(* Logix 5000 project; controller PLC_MCC1300_75F1 vendor 1 type 14 code 166 rev 32.11; software revision 32.04; part 10 of 83 *)

        [35]   // PEG SAMPLE Trailedge Positioning Timer Preset [sec x 100]
        [4].7   // Stress Sample one shot for new LE at Conv 6 Resync Zone
        [6].9   // 400 Deck Conveyor 9 Operate at Trim speed
        [20].3   // STRESS SAMPLE Stop Conv 8 for Sample Positioning
        [32]   // PEG SAMPLE Trailedge Stopping Setpoint [inches x 10]
        [7].8   // PEG SAMPLE Lead-Cap Runout In Progress (Stop Conv 9)
        [50]   // PEG SAMPLE Trailedge Stopping Setpoint [inches x 10]
        [11]   // Sample/Peg CAP Length in Inches
        [7].7   // Sample/Peg Stop Conv 9 When next CAP Arrives
        [37]   // PEG SAMPLE TE Stopping Setpoint for Glass <> 60 In [inches x 10]
        [90]   // PEG SAMPLE Trailedge Stopping(2100in/min) Setpoint [inches x 10]
        [10]   // Sample/Peg CAP Length + Trailedge Position in Zones
        [41]   // 400 DECK Decel Distance for Current Trim Speed [in]
        [2]   // 400 DECK CAP Length of Current Cap [64ths]
        [8]   // Sample/Peg Transfer State Machine
        [14]   // PEG SAMPLE Minimum Gap + Cap Value for LCR [inches / 2]
        [42]   // 400 DECK CAP Length Divided by 2 for Current Piece [in]
        [5].8   // 400 Deck
        [20].2   // Conveyor 7 Leadedge Detected
        [7].2   // Queue Conv 4 Leadedge Detected
        [20].1   // Conveyor 6 Trailedge Detected
        [7].1   // Queue Conv 4 Trailedge Detected
        [0]   // 400 Deck State Variable
        [45]   // 400 Deck Host ID
        [5].9   // 400 Deck
        [25]   // Heavy Glass Sample Cap ID
        [31]   // PEG SAMPLE Decel Distance at Current Speed for Positioning Calc. [in x 10]
        [4].0   // 400 Deck One shot!
   N98 : DINT[40] := ([0] := 12767, [1] := -2664, [5] := 241, [6] := 245, [7] := 244, [8] := 243, [9] := 230, [10] := 232, [11] := 237, [12] := 239);
   O : INT[128] := ([5] := 2#0000_1111_1111_1111, [8] := 2#0000_1000_0000_0000, [9] := 2#0010_0000_0000_1000, [17] := 2#0000_0000_0000_1000, [21] := 2#1111_1100_0000_1000, [23] := 2#0000_0000_0000_0011, [27] := 2#0001_0000_0000_0010, [29] := 2#0001_0000_0000_0010, [30] := 2#0010_0100_0011_1111, [31] := 2#0001_0000_0000_0010, [34] := 2#0000_0000_0000_0110, [38] := 2#0000_0000_0110_0011, [41] := 2#0000_0001_0000_0000, [42] := 2#0000_0000_0000_0100, [46] := 2#0000_0000_0000_0100, [50] := 2#0000_0000_0000_0011, [62] := 2#0000_0000_0000_0011, [66] := 2#0000_0000_0000_0100, [70] := 2#0000_0000_0000_0100, [74] := 2#1000_0100_1100_0011, [78] := 2#0000_0000_0000_0010, [80] := 2#0000_0000_0111_1011, [81] := 2#0000_0010_0100_0000, [82] := 2#0000_0000_0100_0011, [83] := 2#0000_0001_0100_0001, [84] := 2#0000_0001_0100_0001, [85] := 2#0001_0001_0100_0010, [86] := 2#0000_0001_0100_0001, [87] := 2#0001_0000_0000_0010, [89] := 2#0001_0000_0000_0010, [91] := 2#0001_0000_0000_0010, [92] := 2#0000_1001_1100_1010, [93] := 2#0011_0000_0000_0010, [95] := 2#0011_0000_0000_0010, [96] := 2#0000_0000_0000_0011, [97] := 2#0011_0000_0000_0010, [99] := 2#0011_0000_0000_0010, [101] := 2#0011_0001_1100_0010, [103] := 2#0011_0000_0000_0010, [105] := 2#0011_0000_0000_0010, [107] := 2#0011_0000_0000_0010, [109] := 2#0011_0000_0000_0010, [111] := 2#0011_0000_0000_0010, [113] := 2#0011_0000_0000_0010, [115] := 2#0011_0000_0000_0010, [117] := 2#0011_0000_0000_0010, [119] := 2#0011_0000_0000_0010, [121] := 2#0000_0000_1000_0100, [123] := 2#0000_1000_0000_0000);
        [113].8   // VMCC M2 Speed zone 11 Accel Rate Select 1 * M2CM11S
        [113].9   // VMCC M2 Speed zone 11 Accel Rate Select 2 * M2CM11S
        [111].9   // VMCC M2 Speed zone 10 Accel Rate Select 2 * M2CM10N
        [113].10   // VMCC M2 Speed zone 11 Decel Rate Select 1 * M2CM11S
        [103].11   // VMCC M2 Speed zone 8 Decel Rate Select 2 * M2CM8N
        [105].10   // VMCC M2 Speed zone 9 Decel Rate Select 1 * M2CM9S
        [105].11   // VMCC M2 Speed zone 9 Decel Rate Select 2 * M2CM9S
        [107].10   // VMCC M2 Speed zone 9 Decel Rate Select 1 * M2CM9N
        [107].11   // VMCC M2 Speed zone 9 Decel Rate Select 2 * M2CM9N
        [101].2   // VMCC M2 Speed zone 8 Jog * M2CM8S
        [117].6   // VMCC M2 Speed zone 12 Local Control Reques * M2CM12S
        [115].10   // VMCC M2 Speed zone 11 Decel Rate Select 1 * M2CM11N
        [119].4   // VMCC M2 Speed zone 12 Direction Select 1 * M2CM12N
        [119].5   // VMCC M2 Speed zone 12 Direction Select 2 * M2CM12N
        [103].2   // VMCC M2 Speed zone 8 Jog * M2CM8N
        [105].2   // VMCC M2 Speed zone 9 Jog * M2CM9S
        [119].9   // VMCC M2 Speed zone 12 Accel Rate Select 2 * M2CM12N
        [121]   // M2 -->> MB Copy mainline crusher status bits from M2 to MB
        [117].8   // VMCC M2 Speed zone 12 Accel Rate Select 1 * M2CM12S
        [123].2   // M2 -->> MB Trim deck Drive system Critical Failure
        [123].5   // M2 -->> MB Mainline Drive system Critical Failure
        [115].8   // VMCC M2 Speed zone 11 Accel Rate Select 1 * M2CM11N
        [101].3   // VMCC M2 Speed zone 8 Clear Fault * M2CM8S
        [107].2   // VMCC M2 Speed zone 9 Jog * M2CM9N
        [123].11   // M2 -->> MB Drive running M2CM01
        [123].3   // M2 -->> MB Trim deck Drive fault
        [25].3   // ROCKWELL CAPPER Disable auto y-cut bar 4
        [27].0   // VMCC M2 Speed zone 1 Stop * M2CM01
        [5].9   // VMCC M2 Speed zone 10 Foward * 2CM10
        [6].0   // VMCC M2 Speed zone 1 Reverse * 2CM01
        [6].1   // VMCC M2 Speed zone 2 Reverse * 2CM02
        [6].2   // VMCC M2 Speed zone 3 Reverse * 2CM03
        [6].3   // VMCC M2 Speed zone 4 Reverse * 2CM04
        [109].2   // VMCC M2 Speed zone 10 Jog * M2CM10S
        [111].2   // VMCC M2 Speed zone 10 Jog * M2CM10N
        [124].0   // M2 -->> MB Leg 4 Is In Sleep Mode
        [103].3   // VMCC M2 Speed zone 8 Clear Fault * M2CM8N
        [6].4   // VMCC M2 Speed zone 5 Reverse * 2CM05
        [124].1   // M2 -->> MB Leg 5 Is In Sleep Mode
        [6].5   // VMCC M2 Speed zone 6 Reverse * 2CM06
        [123].8   // M2 -->> MB SPARE
        [10].10   // VMCC M2 SPARE
        [10].11   // VMCC M2 SPARE
        [123].9   // M2 -->> MB SPARE
        [20].8   // VMCC TD Trim knocker Speed select 2
        [124].4   // M2-->MB VISION SYS Rejected Plate Alarm Horn
        [19].2   // VMCC TD Trim Zone 1 North knocker Adjust motor
        [105].3   // VMCC M2 Speed zone 9 Clear Fault * M2CM9S
        [113].2   // VMCC M2 Speed zone 11 Jog * M2CM11S
        [107].3   // VMCC M2 Speed zone 9 Clear Fault * M2CM9N
        [123].13   // M2 -->> MB Crush-all Selector sw. Status
        [20].9   // VMCC TD Trim deck Speed select 2 North side
        [101].12   // VMCC M2 Speed zone 8 Speed Select 1 * M2CM8S
        [42].5   // RELIANCE CAPPING SYSTEM Tracking window Lamp
        [19].3   // VMCC TD Trim Zone 1 South knocker Adjust motor
        [70].5   // RELIANCE CAPPING SYSTEM Tracking window Lamp
        [115].2   // VMCC M2 Speed zone 11 Jog * M2CM11N
        [19].4   // VMCC TD Trim Zone 2 North knocker Adjust motor
        [19].5   // VMCC TD Trim Zone 2 South knocker Adjust motor
        [27].3   // VMCC M2 Speed zone 1 Clear Fault * M2CM01
        [7].10   // VMCC M2 Speed zone 11 Speed Select 2 * 2CM11
        [22].2   // VMCC TD Trim Zone 1 North trim Adjust motor
        [22].3   // VMCC TD Trim Zone 1 South trim Adjust motor
        [117].9   // VMCC M2 Speed zone 12 Accel Rate Select 2 * M2CM12S
        [74].13   // BENCHBOARD SPARE
        [101].13   // VMCC M2 Speed zone 8 Speed Select 2 * M2CM8S
        [109].10   // VMCC M2 Speed zone 10 Decel Rate Select 1 * M2CM10S
        [109].11   // VMCC M2 Speed zone 10 Decel Rate Select 2 * M2CM10S
        [109].6   // VMCC M2 Speed zone 10 Local Control Reques * M2CM10S
        [109].8   // VMCC M2 Speed zone 10 Accel Rate Select 1 * M2CM10S
        [25].4   // ROCKWELL CAPPER Disable auto y-cut bar 3
        [10].12   // VMCC M2 SPARE
        [10].13   // VMCC M2 SPARE
        [10].14   // VMCC M2 SPARE
        [10].15   // VMCC M2 SPARE
        [19].12   // VMCC TD SPARE
        [19].13   // VMCC TD SPARE
        [19].14   // VMCC TD SPARE
        [19].15   // VMCC TD SPARE
        [101].0   // VMCC M2 Speed zone 8 Stop * M2CM8S
        [19].6   // VMCC TD Trim Zone 3 North knocker Adjust motor
        [125]   // MB -->> M2 Host comp. Reliance Crossbreaks Disable Ycuts
        [119].6   // VMCC M2 Speed zone 12 Local Control Reques * M2CM12N
        [109].0   // VMCC M2 Speed zone 10 Stop * M2CM10S
        [111].0   // VMCC M2 Speed zone 10 Stop * M2CM10N
        [113].0   // VMCC M2 Speed zone 11 Stop * M2CM11S
        [115].0   // VMCC M2 Speed zone 11 Stop * M2CM11N
        [42].2   // PANEL TD-CS2N North Trim knocker #2 Lower
        [46].2   // PANEL TD-CS3N North Trim knocker #3 Lower
        [50].2   // PANEL TD-CS4N North Trim knocker #4 Lower
        [55].2   // PANEL TD-CS5N North Trim knocker #5 Lower
        [62].2   // PANEL TD-CS4S South Trim knocker #4 Lower
        [66].2   // PANEL TD-CS3S South Trim knocker #3 Lower
        [70].2   // PANEL TD-CS2S South Trim knocker #2 Lower
        [7].0   // VMCC M2 Speed zone 1 Speed Select 2 * 2CM01
        [7].1   // VMCC M2 Speed zone 2 Speed Select 2 * 2CM02
        [7].2   // VMCC M2 Speed zone 3 Speed Select 2 * 2CM03
        [7].3   // VMCC M2 Speed zone 4 Speed Select 2 * 2CM04
        [7].4   // VMCC M2 Speed zone 5 Speed Select 2 * 2CM05
        [7].5   // VMCC M2 Speed zone 6 Speed Select 2 * 2CM06
        [7].6   // VMCC M2 Speed zone 7 Speed Select 2 * 2CM07
        [7].7   // VMCC M2 Speed zone 8 Speed Select 2 * 2CM08
        [7].8   // VMCC M2 Speed zone 9 Speed Select 2 * 2CM09
        [85].3   // VMCC M2 Speed zone 4 Clear Fault * M2CM4S
        [87].3   // VMCC M2 Speed zone 4 Clear Fault * M2CM4N
        [22].0   // VMCC TD Krurl drop North trim Adjust motor
        [89].3   // VMCC M2 Speed zone 5 Clear Fault * M2CM5S
        [8].0   // VMCC M2 Speed zone 1 Speed Select 1 * 2CM01
        [8].1   // VMCC M2 Speed zone 2 Speed Select 1 * 2CM02
        [8].2   // VMCC M2 Speed zone 3 Speed Select 1 * 2CM03
        [8].3   // VMCC M2 Speed zone 4 Speed Select 1 * 2CM04
        [8].4   // VMCC M2 Speed zone 5 Speed Select 1 * 2CM05
        [8].5   // VMCC M2 Speed zone 6 Speed Select 1 * 2CM06
        [8].6   // VMCC M2 Speed zone 7 Speed Select 1 * 2CM07
        [8].7   // VMCC M2 Speed zone 8 Speed Select 1 * 2CM08
        [22].1   // VMCC TD Krurl drop South trim Adjust motor
        [25].1   // ROCKWELL CAPPER Disable manual y-cut bar 2
        [8].8   // VMCC M2 Speed zone 9 Speed Select 1 * 2CM09
        [25].5   // ROCKWELL CAPPER Disable auto y-cut bar 2
        [103].0   // VMCC M2 Speed zone 8 Stop * M2CM8N
        [117].0   // VMCC M2 Speed zone 12 Stop * M2CM12S
        [119].0   // VMCC M2 Speed zone 12 Stop * M2CM12N
        [105].0   // VMCC M2 Speed zone 9 Stop * M2CM9S
        [115].11   // VMCC M2 Speed zone 11 Decel Rate Select 2 * M2CM11N
        [91].3   // VMCC M2 Speed zone 5 Clear Fault * M2CM5N
        [117].2   // VMCC M2 Speed zone 12 Jog * M2CM12S
        [119].2   // VMCC M2 Speed zone 12 Jog * M2CM12N
        [123].14   // M2 -->> MB Leg 2 Is In Sleep Mode
        [123].15   // M2 -->> MB Leg 3 Is In Sleep Mode
        [22].4   // VMCC TD Trim Zone 2 North trim Adjust motor
        [20].12   // VMCC TD Trim knocker Speed select 1
        [6].10   // VMCC M2 Speed zone 11 Reverse * 2CM11
        [6].11   // VMCC M2 Speed zone 12 Reverse * 2CM12
        [9].2   // VMCC M2 SPARE
        [123].10   // M2 -->> MB SPARE
        [10].0   // VMCC M2 SPARE
        [22].5   // VMCC TD Trim Zone 2 South trim Adjust motor
        [22].6   // VMCC TD Trim Zone 3 North trim Adjust motor
        [101].14   // VMCC M2 Speed zone 8 Speed Select 3 * M2CM8S
        [103].12   // VMCC M2 Speed zone 8 Speed Select 1 * M2CM8N
        [8].10   // VMCC M2 Speed zone 11 Speed Select 1 * 2CM11
        [19].7   // VMCC TD Trim Zone 3 South knocker Adjust motor
        [8].11   // VMCC M2 Speed zone 12 Speed Select 1 * 2CM12
        [103].13   // VMCC M2 Speed zone 8 Speed Select 2 * M2CM8N
        [19]   // TRIM KNOCKERS Contactors used For drive to Knocker adj Motors
        [119].8   // VMCC M2 Speed zone 12 Accel Rate Select 1 * M2CM12N
        [22].7   // VMCC TD Trim Zone 3 South trim Adjust motor
        [22].8   // VMCC TD Trim Zone 4 North trim Adjust motor
        [103].14   // VMCC M2 Speed zone 8 Speed Select 3 * M2CM8N
        [105].12   // VMCC M2 Speed zone 9 Speed Select 1 * M2CM9S
        [93].3   // VMCC M2 Speed zone 6 Clear Fault * M2CM6S
        [22].9   // VMCC TD Trim Zone 4 South trim Adjust motor
        [27].1   // VMCC M2 Speed zone 1 Forward/start * M2CM01
        [19].8   // VMCC TD Trim Zone 4 North knocker Adjust motor
        [105].13   // VMCC M2 Speed zone 9 Speed Select 2 * M2CM9S
        [115].4   // VMCC M2 Speed zone 11 Direction Select 1 * M2CM11N
        [19].9   // VMCC TD Trim Zone 4 South knocker Adjust motor
        [95].3   // VMCC M2 Speed zone 6 Clear Fault * M2CM6N
        [105].14   // VMCC M2 Speed zone 9 Speed Select 3 * M2CM9S
        [115].9   // VMCC M2 Speed zone 11 Accel Rate Select 2 * M2CM11N
        [25].6   // ROCKWELL CAPPER Disable auto y-cut bar 1
        [29].3   // VMCC M2 Speed zone 2 Clear Fault * M2CM2
        [31].3   // VMCC M2 Speed zone 3 Clear Fault * M2CM3
        [38].3   // PANEL TD-CS1N North Trim knocker 1 Lower
        [27].13   // VMCC M2 Speed zone 1 Speed Select 1 * M2CM01
        [82].3   // PANEL TD-CS1S South Trim knocker 1 Lower
        [6].6   // VMCC M2 Speed zone 7 Reverse * 2CM07
        [25].2   // ROCKWELL CAPPER Disable manual y-cut bar 1
        [6].9   // VMCC M2 Speed zone 10 Reverse * 2CM10
        [85].1   // VMCC M2 Speed zone 4 Forward/start * M2CM4S
        [115].5   // VMCC M2 Speed zone 11 Direction Select 2 * M2CM11N
        [87].1   // VMCC M2 Speed zone 4 Forward/start * M2CM4N
        [25].0   // ROCKWELL CAPPER Crossbreak in progress
        [54].3   // PANEL TD-CS5N Reject window Lamp North
        [58].3   // PANEL TD-CS5S Reject window Lamp South
        [38].4   // Trim Deck Float Glass Hold Down Wheel Solenoid
        [89].1   // VMCC M2 Speed zone 5 Forward/start * M2CM5S
        [107].12   // VMCC M2 Speed zone 9 Speed Select 1 * M2CM9N
        [107].13   // VMCC M2 Speed zone 9 Speed Select 2 * M2CM9N
        [107].14   // VMCC M2 Speed zone 9 Speed Select 3 * M2CM9N
        [19].10   // VMCC TD Trim Zone 5 North knocker Adjust motor
        [19].11   // VMCC TD Trim Zone 5 South knocker Adjust motor
        [34].0   // PANEL KD-CS1N North Knurl knocker Auto mode Lamp
        [9].4   // VMCC M2 Red Stack lite
        [97].3   // VMCC M2 Speed zone 7 Clear Fault * M2CM7S
        [29].1   // VMCC M2 Speed zone 2 Forward/start * M2CM2
        [109].9   // VMCC M2 Speed zone 10 Accel Rate Select 2 * M2CM10S
        [111].10   // VMCC M2 Speed zone 10 Decel Rate Select 1 * M2CM10N
        [99].3   // VMCC M2 Speed zone 7 Clear Fault * M2CM7N
        [109].15   // VMCC M2 Speed zone 10 MOP Decrement * M2CM10S
        [111].15   // VMCC M2 Speed zone 10 MOP Decrement * M2CM10N
        [113].15   // VMCC M2 Speed zone 11 MOP Decrement * M2CM11S
        [115].15   // VMCC M2 Speed zone 11 MOP Decrement * M2CM11N
        [117].15   // VMCC M2 Speed zone 12 MOP Decrement * M2CM12S
        [119].15   // VMCC M2 Speed zone 12 MOP Decrement * M2CM12N
        [38].0   // PANEL TD-CS1N North Trim knocker 1 Auto mode Lamp
        [38].1   // PANEL TD-CS1N South Trim knocker 1 Auto mode Lamp
        [38].6   // Float Glass Hold Down Wheels Up Manual Oper. Lamp
        [123].0   // M2 -->> MB Drop #1 Crusher Pushbutton
        [34].2   // PANEL KD-CS1N North Knurl knocker Lower
        [74].10   // BENCHBOARD Knurl Nth & Sth Auto Mode
        [78].2   // PANEL KD-CS1S South Knurl knocker Lower
        [117].10   // VMCC M2 Speed zone 12 Decel Rate Select 1 * M2CM12S
        [117].11   // VMCC M2 Speed zone 12 Decel Rate Select 2 * M2CM12S
        [46].3   // Trim Deck PANEL TD-CS3N Crush all Switch Pilot Light
        [66].3   // Trim Deck PANEL TD-CS3S Crush all Switch Pilot Light
        [82].0   // PANEL TD-CS1S North Trim knocker 1 Auto mode Lamp
        [34].1   // PANEL KD-CS1N South Knurl knocker Auto mode Lamp
        [78].0   // PANEL KD-CS1S North Knurl knocker Auto mode Lamp
        [31].1   // VMCC M2 Speed zone 3 Forward/start * M2CM3
        [38].5   // Trim Deck Eclipse Hold Down Wheel Solenoid
        [38].7   // Eclipse Hold Down Wheels Manual Oper. Lamp
        [5]   // Word containing Drive forward Bits for Conveyors
        [7].9   // VMCC M2 Speed zone 10 Speed Select 2 * 2CM10
        [82].7   // Eclipse Hold Down Wheels Manual Oper. Lamp
        [8].9   // VMCC M2 Speed zone 10 Speed Select 1 * 2CM10
        [78].1   // PANEL KD-CS1S South Knurl knocker Auto mode Lamp
        [7].11   // VMCC M2 Speed zone 12 Ref Speed\\Select 3 2CM12N
        [113].11   // VMCC M2 Speed zone 11 Decel Rate Select 2 * M2CM11S
        [119].10   // VMCC M2 Speed zone 12 Decel Rate Select 1 * M2CM12N
        [119].11   // VMCC M2 Speed zone 12 Decel Rate Select 2 * M2CM12N
        [117].4   // VMCC M2 Speed zone 12 Direction Select 1 * M2CM12S
        [117].5   // VMCC M2 Speed zone 12 Direction Select 2 * M2CM12S
        [113].5   // VMCC M2 Speed zone 11 Direction Select 2 * M2CM11S
        [113].6   // VMCC M2 Speed zone 11 Local Control Reques * M2CM11S
        [82].1   // PANEL TD-CS1S South Trim knocker 1 Auto mode Lamp
        [107].0   // VMCC M2 Speed zone 9 Stop * M2CM9N
        [101].4   // VMCC M2 Speed zone 8 Direction Select 1 * M2CM8S
        [115].6   // VMCC M2 Speed zone 11 Local Control Reques * M2CM11N
        [101].5   // VMCC M2 Speed zone 8 Direction Select 2 * M2CM8S
        [82].6   // Float Glass Hold Down Wheels Manual Oper. Lamp
        [85].12   // VMCC M2 Speed zone 4 Speed Select 1 * M2CM4S
        [85].13   // VMCC M2 Speed zone 4 Speed Select 2 * M2CM4S
        [87].12   // VMCC M2 Speed zone 4 Speed Select 1 * M2CM4N
        [87].13   // VMCC M2 Speed zone 4 Speed Select 2 * M2CM4N
        [89].12   // VMCC M2 Speed zone 5 Speed Select 1 * M2CM5S
        [89].13   // VMCC M2 Speed zone 5 Speed Select 2 * M2CM5S
        [91].12   // VMCC M2 Speed zone 5 Speed Select 1 * M2CM5N
        [91].13   // VMCC M2 Speed zone 5 Speed Select 2 * M2CM5N
        [93].12   // VMCC M2 Speed zone 6 Speed Select 1 * M2CM6S
        [93].13   // VMCC M2 Speed zone 6 Speed Select 2 * M2CM6S
        [95].12   // VMCC M2 Speed zone 6 Speed Select 1 * M2CM6N
        [95].13   // VMCC M2 Speed zone 6 Speed Select 2 * M2CM6N
        [97].12   // VMCC M2 Speed zone 7 Speed Select 1 * M2CM7S
        [111].11   // VMCC M2 Speed zone 10 Decel Rate Select 2 * M2CM10N
        [111].6   // VMCC M2 Speed zone 10 Local Control Reques * M2CM10N
        [111].8   // VMCC M2 Speed zone 10 Accel Rate Select 1 * M2CM10N
        [97].13   // VMCC M2 Speed zone 7 Speed Select 2 * M2CM7S
        [99].12   // VMCC M2 Speed zone 7 Speed Select 1 * M2CM7N
        [99].13   // VMCC M2 Speed zone 7 Speed Select 2 * M2CM7N
        [101].15   // VMCC M2 Speed zone 8 MOP Decrement * M2CM8S
        [103].15   // VMCC M2 Speed zone 8 MOP Decrement * M2CM8N
        [105].15   // VMCC M2 Speed zone 9 MOP Decrement * M2CM9S
        [107].15   // VMCC M2 Speed zone 9 MOP Decrement * M2CM9N
        [109].1   // VMCC M2 Speed zone 10 Forward/start * M2CM10S
        [101].1   // VMCC M2 Speed zone 8 Forward/start * M2CM8S
        [101].7   // VMCC M2 Speed zone 8 MOP Increment * M2CM8S
        [103].1   // VMCC M2 Speed zone 8 Forward/start * M2CM8N
        [103].7   // VMCC M2 Speed zone 8 MOP Increment * M2CM8N
        [105].1   // VMCC M2 Speed zone 9 Forward/start * M2CM9S
        [105].7   // VMCC M2 Speed zone 9 MOP Increment * M2CM9S
        [107].1   // VMCC M2 Speed zone 9 Forward/start * M2CM9N
        [103].4   // VMCC M2 Speed zone 8 Direction Select 1 * M2CM8N
        [103].5   // VMCC M2 Speed zone 8 Direction Select 2 * M2CM8N
        [20].1   // VMCC TD Trim deck Forward North side
        [20].2   // VMCC TD Trim deck Forward South side
        [20].5   // VMCC TD Trim deck Reverse North side
        [20].6   // VMCC TD Trim deck Reverse South side
        [5].10   // VMCC M2 Speed zone 11 Foward * 2CM11
        [5].11   // VMCC M2 Speed zone 12 Foward * 2CM12
        [74].12   // BENCHBOARD Crossbreak Alert Buzzer
        [123].1   // M2 -->> MB Trim deck E-stop
        [123].12   // M2 -->> MB Mainline Backup to
        [123].4   // M2 -->> MB Mainline E-stop
        [123].6   // M2 -->> MB Mainline Drive fault
        [124].2   // M2 -->> MB ML Is In Sleep Mode
        [124].3   // M2-->MB UL Crusher Is Faulted
        [127].4   // M2-->MB Float Glass Prodution
        [20].0   // VMCC TD Trim knocker Forward
        [20].4   // VMCC TD Trim knocker Reverse
        [21].0   // VMCC TD Drive fault Lamp
        [21].1   // VMCC TD Drive fault Reset relay
        [21].3   // VMCC TD Alarm horn Relay
        [107].7   // VMCC M2 Speed zone 9 MOP Increment * M2CM9N
        [109].3   // VMCC M2 Speed zone 10 Clear Fault * M2CM10S
        [109].7   // VMCC M2 Speed zone 10 MOP Increment * M2CM10S
        [111].1   // VMCC M2 Speed zone 10 Forward/start * M2CM10N
        [111].7   // VMCC M2 Speed zone 10 MOP Increment * M2CM10N
        [113].1   // VMCC M2 Speed zone 11 Forward/start * M2CM11S
        [113].7   // VMCC M2 Speed zone 11 MOP Increment * M2CM11S
        [115].1   // VMCC M2 Speed zone 11 Forward/start * M2CM11N
        [111].3   // VMCC M2 Speed zone 10 Clear Fault * M2CM10N
        [113].3   // VMCC M2 Speed zone 11 Clear Fault * M2CM11S
        [115].3   // VMCC M2 Speed zone 11 Clear Fault * M2CM11N
        [117].3   // VMCC M2 Speed zone 12 Clear Fault * M2CM12S
        [119].3   // VMCC M2 Speed zone 12 Clear Fault * M2CM12N
        [19].0   // VMCC TD Krurl drop North knocker Adjust motor
        [19].1   // VMCC TD Krurl drop South knocker Adjust motor
        [20].10   // VMCC TD Trim deck Speed select 2 South side
        [20].13   // VMCC TD Trim deck Speed select 1 North side
        [20].14   // VMCC TD Trim deck Speed select 1 South side
        [115].7   // VMCC M2 Speed zone 11 MOP Increment * M2CM11N
        [117].1   // VMCC M2 Speed zone 12 Forward/start * M2CM12S
        [117].7   // VMCC M2 Speed zone 12 MOP Increment * M2CM12S
        [119].1   // VMCC M2 Speed zone 12 Forward/start * M2CM12N
        [22].10   // VMCC TD Trim Zone 5 North trim Adjust motor
        [22].11   // VMCC TD Trim Zone 5 South trim Adjust motor
        [27].12   // VMCC M2 Speed zone 1 Speed Select 1 * M2CM1
        [29].12   // VMCC M2 Speed zone 2 Speed Select 1 * M2CM2
        [29].13   // VMCC M2 Speed zone 2 Speed Select 2 * M2CM2
        [31].12   // VMCC M2 Speed zone 3 Speed Select 1 * M2CM3
        [31].13   // VMCC M2 Speed zone 3 Speed Select 2 * M2CM3
        [91].1   // VMCC M2 Speed zone 5 Forward/start * M2CM5N
        [93].1   // VMCC M2 Speed zone 6 Forward/start * M2CM6S
        [95].1   // VMCC M2 Speed zone 6 Forward/start * M2CM6N
        [97].1   // VMCC M2 Speed zone 7 Forward/start * M2CM7S
        [20].11   // VMCC TD SPARE
        [20].15   // VMCC TD SPARE
        [21].10   // VMCC TD SPARE
        [9].7   // VMCC M2 SPARE
        [9].8   // VMCC M2 SPARE
        [21].4   // VMCC TD Red Stack lite
        [21].5   // VMCC TD Blue Stack lite
        [6].7   // VMCC M2 Speed zone 8 Reverse * 2CM08
        [6].8   // VMCC M2 Speed zone 9 Reverse * 2CM09
        [119].7   // VMCC M2 Speed zone 12 MOP Increment * M2CM12N
        [99].1   // VMCC M2 Speed zone 7 Forward/start * M2CM7N
        [105].4   // VMCC M2 Speed zone 9 Direction Select 1 * M2CM9S
        [105].5   // VMCC M2 Speed zone 9 Direction Select 2 * M2CM9S
        [54].2   // PANEL TD-CS5N Reliance data Received Lamp North
        [107].4   // VMCC M2 Speed zone 9 Direction Select 1 * M2CM9N
        [107].5   // VMCC M2 Speed zone 9 Direction Select 2 * M2CM9N
        [58].2   // PANEL TD-CS5S Reliance Data received Lamp South
        [109].12   // VMCC M2 Speed zone 10 Speed Select 1 * M2CM10S
        [109].13   // VMCC M2 Speed zone 10 Speed Select 2 * M2CM10S
        [109].14   // VMCC M2 Speed zone 10 Speed Select 3 * M2CM10S
        [111].12   // VMCC M2 Speed zone 10 Speed Select 1 * M2CM10N
        [101].8   // VMCC M2 Speed zone 8 Accel Rate Select 1 * M2CM8S
        [111].13   // VMCC M2 Speed zone 10 Speed Select 2 * M2CM10N
        [111].14   // VMCC M2 Speed zone 10 Speed Select 3 * M2CM10N
        [113].12   // VMCC M2 Speed zone 11 Speed Select 1 * M2CM11S
        [101].6   // VMCC M2 Speed zone 8 Local Control Reques * M2CM8S
        [103].6   // VMCC M2 Speed zone 8 Local Control Reques * M2CM8N
        [10].1   // VMCC M2 SPARE
        [10].2   // VMCC M2 SPARE
        [21].11   // VMCC TD SPARE
        [21].12   // VMCC TD SPARE
        [21].13   // VMCC TD SPARE
        [21].14   // VMCC TD SPARE
        [21].15   // VMCC TD SPARE
        [22].12   // VMCC TD SPARE
        [10].3   // VMCC M2 SPARE
        [10].4   // VMCC M2 SPARE
        [10].5   // VMCC M2 SPARE
        [10].6   // VMCC M2 SPARE
        [10].7   // VMCC M2 SPARE
        [10].8   // VMCC M2 SPARE
        [10].9   // VMCC M2 SPARE
        [20].3   // VMCC TD SPARE
        [113].13   // VMCC M2 Speed zone 11 Speed Select 2 * M2CM11S
        [113].14   // VMCC M2 Speed zone 11 Speed Select 3 * M2CM11S
        [115].12   // VMCC M2 Speed zone 11 Speed Select 1 * M2CM11N
        [103].8   // VMCC M2 Speed zone 8 Accel Rate Select 1 * M2CM8N
        [103].9   // VMCC M2 Speed zone 8 Accel Rate Select 2 * M2CM8N
        [115].13   // VMCC M2 Speed zone 11 Speed Select 2 * M2CM11N
        [115].14   // VMCC M2 Speed zone 11 Speed Select 3 * M2CM11N
        [117].12   // VMCC M2 Speed zone 12 Speed Select 1 * M2CM12S
        [105].6   // VMCC M2 Speed zone 9 Local Control Reques * M2CM9S
        [105].8   // VMCC M2 Speed zone 9 Accel Rate Select 1 * M2CM9S
        [117].13   // VMCC M2 Speed zone 12 Speed Select 2 * M2CM12S
        [117].14   // VMCC M2 Speed zone 12 Speed Select 3 * M2CM12S
        [119].12   // VMCC M2 Speed zone 12 Speed Select 1 * M2CM12N
        [105].9   // VMCC M2 Speed zone 9 Accel Rate Select 2 * M2CM9S
        [107].6   // VMCC M2 Speed zone 9 Local Control Reques * M2CM9N
        [119].13   // VMCC M2 Speed zone 12 Speed Select 2 * M2CM12N
        [119].14   // VMCC M2 Speed zone 12 Speed Select 3 * M2CM12N
        [42].0   // PANEL TD-CS2N North Trim knocker #2 Auto mode Lamp
        [107].8   // VMCC M2 Speed zone 9 Accel Rate Select 1 * M2CM9N
        [107].9   // VMCC M2 Speed zone 9 Accel Rate Select 2 * M2CM9N
        [101].10   // VMCC M2 Speed zone 8 Decel Rate Select 1 * M2CM8S
        [42].1   // PANEL TD-CS2N South Trim knocker #2 Auto mode Lamp
        [46].0   // PANEL TD-CS3N North Trim knocker #3 Auto mode Lamp
        [46].1   // PANEL TD-CS3N South Trim knocker #3 Auto mode Lamp
        [109].4   // VMCC M2 Speed zone 10 Direction Select 1 * M2CM10S
        [109].5   // VMCC M2 Speed zone 10 Direction Select 2 * M2CM10S
        [101].11   // VMCC M2 Speed zone 8 Decel Rate Select 2 * M2CM8S
        [21].6   // VMCC TD Amber Stack lite
        [111].4   // VMCC M2 Speed zone 10 Direction Select 1 * M2CM10N
        [74].0   // BENCHBOARD Trim #1 North Auto mode
        [101].9   // VMCC M2 Speed zone 8 Accel Rate Select 2 * M2CM8S
        [29].0   // VMCC M2 Speed zone 2 Stop * M2CM2
        [103].10   // VMCC M2 Speed zone 8 Decel Rate Select 1 * M2CM8N
        [22].13   // VMCC TD SPARE
        [22].14   // VMCC TD SPARE
        [22].15   // VMCC TD SPARE
        [20].7   // VMCC TD SPARE
        [21].2   // VMCC TD SPARE
        [21].7   // VMCC TD SPARE
        [21].8   // VMCC TD SPARE
        [21].9   // VMCC TD SPARE
        [5].12   // VMCC M2 SPARE
        [74].1   // BENCHBOARD Trim #1 South Auto mode
        [31].0   // VMCC M2 Speed zone 3 Stop * M2CM3
        [38].2   // PANEL TD-CS1N Snap roll Extend
        [50].0   // PANEL TD-CS4N North Trim knocker #4 Auto mode Lamp
        [50].1   // PANEL TD-CS4N South Trim knocker #4 Auto mode Lamp
        [54].0   // PANEL TD-CS5N North Trim knocker #5 Auto mode Lamp
        [54].1   // PANEL TD-CS5N South Trim knocker #5 Auto mode Lamp
        [111].5   // VMCC M2 Speed zone 10 Direction Select 2 * M2CM10N
        [55].0   // PANEL TD-CS5N North Trim knocker #5 Auto mode Lamp
        [55].1   // PANEL TD-CS5N South Trim knocker #5 Auto mode Lamp
        [58].0   // PANEL TD-CS5S North Trim knocker #5 Auto mode Lamp
        [58].1   // PANEL TD-CS5S South Trim knocker #5 Auto mode Lamp
        [62].0   // PANEL TD-CS4S North Trim knocker #4 Auto mode Lamp
        [62].1   // PANEL TD-CS4S South Trim knocker #4 Auto mode Lamp
        [66].0   // PANEL TD-CS3S North Trim knocker #3 Auto mode Lamp
        [66].1   // PANEL TD-CS3S South Trim knocker #3 Auto mode Lamp
        [5].0   // VMCC M2 Speed zone 1 Foward * 2CM01
        [5].1   // VMCC M2 Speed zone 2 Foward * 2CM02
        [5].13   // VMCC M2 SPARE
        [5].14   // VMCC M2 SPARE
        [5].15   // VMCC M2 SPARE
        [6].12   // VMCC M2 SPARE
        [5].2   // VMCC M2 Speed zone 3 Foward * 2CM03
        [5].3   // VMCC M2 Speed zone 4 Foward * 2CM04
        [5].4   // VMCC M2 Speed zone 5 Foward * 2CM05
        [5].5   // VMCC M2 Speed zone 6 Foward * 2CM06
        [5].6   // VMCC M2 Speed zone 7 Foward * 2CM07
        [5].7   // VMCC M2 Speed zone 8 Foward * 2CM08
        [5].8   // VMCC M2 Speed zone 9 Foward * 2CM09
        [74].11   // BENCHBOARD Trim master
        [70].0   // PANEL TD-CS2S North Trim knocker #2 Auto mode Lamp
        [70].1   // PANEL TD-CS2S South Trim knocker #2 Auto mode Lamp
        [74].14   // Reliance BENCHBOARD Crush all Switch Pilot Light
        [113].4   // VMCC M2 Speed zone 11 Direction Select 1 * M2CM11S
        [74].15   // BENCHBOARD No. 1 crusher Down
        [74].2   // BENCHBOARD Trim #2 North Auto mode
        [6].13   // VMCC M2 SPARE
        [6].14   // VMCC M2 SPARE
        [6].15   // VMCC M2 SPARE
        [7].12   // VMCC M2 SPARE
        [74].3   // BENCHBOARD Trim #2 South Auto mode
        [74].4   // BENCHBOARD Trim #3 North Auto mode
        [74].5   // BENCHBOARD Trim #3 South Auto mode
        [74].6   // BENCHBOARD Trim #4 North Auto mode
        [74].7   // BENCHBOARD Trim #4 South Auto mode
        [74].8   // BENCHBOARD Trim #5 North Auto mode
        [74].9   // BENCHBOARD Trim #5 South Auto mode
        [82].2   // PANEL TD-CS1S Snap roll Extend
        [85].0   // VMCC M2 Speed zone 4 Stop * M2CM4S
        [87].0   // VMCC M2 Speed zone 4 Stop * M2CM4N
        [89].0   // VMCC M2 Speed zone 5 Stop * M2CM5S
        [91].0   // VMCC M2 Speed zone 5 Stop * M2CM5N
        [93].0   // VMCC M2 Speed zone 6 Stop * M2CM6S
        [95].0   // VMCC M2 Speed zone 6 Stop * M2CM6N
        [97].0   // VMCC M2 Speed zone 7 Stop * M2CM7S
        [99].0   // VMCC M2 Speed zone 7 Stop * M2CM7N
        [9].0   // VMCC M2 Drive fault Lamp
        [7].13   // VMCC M2 SPARE
        [7].14   // VMCC M2 SPARE
        [7].15   // VMCC M2 SPARE
        [8].12   // VMCC M2 SPARE
        [82].15   // VMCC M2 Speed zone 1 speed up signal Indicator Light for Snap Roll Camera
        [9].1   // VMCC M2 Drive fault Reset relay
        [9].3   // VMCC M2 Alarm horn Relay
        [9].5   // VMCC M2 Blue Stack lite
        [8].13   // VMCC M2 SPARE
        [8].14   // VMCC M2 SPARE
        [8].15   // VMCC M2 SPARE
        [9].10   // VMCC M2 SPARE
        [9].6   // VMCC M2 Amber Stack lite
        [9].11   // VMCC M2 SPARE
        [9].12   // VMCC M2 SPARE
        [9].13   // VMCC M2 SPARE
        [9].14   // VMCC M2 SPARE
        [9].15   // VMCC M2 SPARE
        [9].9   // VMCC M2 SPARE
   QC1_RES_LMP : ALIAS FOR O[36].2;
   QC2_PE_N : ALIAS FOR B3[12].15;
   QC2_PE_S : ALIAS FOR I[36].3;
   QC2_PE_SOUTH : ALIAS FOR B3[6].11;
   QC2_RES_LMP : ALIAS FOR O[36].3;
   QC3_PE : ALIAS FOR B3[6].12;
   QC3_PE_N : ALIAS FOR B3[13].0;
   QC3_PE_S : ALIAS FOR I[36].4;
   QC3_RES_LMP : ALIAS FOR O[36].4;
   QC4_LE_DET : ALIAS FOR N95[7].2;
   QC4_PE_N : ALIAS FOR B3[13].1;
   QC4_PE_S : ALIAS FOR B3[6].13;
   QC4_RES_LMP : ALIAS FOR O[36].5;
   QC4_TE_DET : ALIAS FOR N95[7].1;
   QC5_PE_N : ALIAS FOR B3[13].2;
   QC5_PE_S : ALIAS FOR B3[6].14;
   QC5_RES_LMP : ALIAS FOR O[36].6;
   QC6_PE_S : ALIAS FOR I[10].5;
   R150 : CONTROL[1];
   R186 : CONTROL[1];
   R19 : CONTROL[4] := ([1].LEN := 12, [2].LEN := 12);
        [1]   // MOTOR SPEED CALCULATION FAL control block
   R19_001_POS : ALIAS FOR R19[1].POS;
   R19_002_POS : ALIAS FOR R19[2].POS;
   R509 : CONTROL[4] := ([0].LEN := 12, [0].POS := 11, [0].EN := 1, [0].DN := 1, [1].LEN := 1, [1].EN := 1, [1].DN := 1, [2].LEN := 12, [3].LEN := 1, [3].EN := 1, [3].DN := 1);
        [0].DN   // MOTOR SPEED CALCULATION FAL control Error bit
        [0].ER   // MOTOR SPEED CALCULATION FAL control Error bit
        [0]   // MOTOR SPEED CALCULATION FAL control block
        [1]   // MOTOR SPEED CALCULATION FAL control block